screen "分段捻缩" 1280x740, template "模板_设置"
   on GenerateScreen: "TitleUpdater"()
   TextField "Text Field_41" at 427,24 size 154x42; Text '分段捻缩'
   TextField "Text Field_48" at 136,126 size 119x56; Text '第一段:'
   TextField "Text Field_49" at 800,124 size 84x56; Text 'mm/s'
   IOField "IO Field_56" at 693,124 size 91x56; FormatPattern 99.9
      ProcessValue <- "ST_VAR_ZhangLi_HMI_r64Velocity_NianSuo_n{0}"
   IOField "IO Field_1" at 257,126 size 94x56; FormatPattern 999
      ProcessValue <- "ST_VAR_ZhangLi_HMI_r64NianDu_NianSuo_Percent_n{0}"
   TextField "Text Field_2" at 349,125 size 117x56; Text '% ～'
   IOField "IO Field_2" at 440,124 size 115x56; FormatPattern 99.9
      ProcessValue <- "ST_VAR_ZhangLi_HMI_r64NianDu_NianSuo_Percent_n{1}"
   TextField "Text Field_3" at 557,124 size 60x56; Text '%,'
   TextField "Text Field_4" at 604,124 size 82x56; Text '速度:'
   IOField "IO Field_3" at 257,194 size 92x56; FormatPattern 9999
      ProcessValue <- "ST_VAR_ZhangLi_HMI_r64NianDu_NianSuo_n{0}"
   IOField "IO Field_4" at 440,190 size 115x56; FormatPattern 9999
      ProcessValue <- "ST_VAR_ZhangLi_HMI_r64NianDu_NianSuo_n{1}"
   TextField "Text Field_5" at 349,194 size 82x56; Text '捻～'
   TextField "Text Field_6" at 558,190 size 82x56; Text '捻'
   TextField "Text Field_1" at 134,279 size 119x56; Text '第二段:'
   TextField "Text Field_7" at 798,277 size 84x56; Text 'mm/s'
   IOField "IO Field_5" at 691,277 size 91x56; FormatPattern 99.9
      ProcessValue <- "ST_VAR_ZhangLi_HMI_r64Velocity_NianSuo_n{1}"
   IOField "IO Field_6" at 255,279 size 94x56; FormatPattern 99.9
      ProcessValue <- "ST_VAR_ZhangLi_HMI_r64NianDu_NianSuo_Percent_n{1}"
   TextField "Text Field_8" at 347,278 size 117x56; Text '% ～'
   IOField "IO Field_7" at 438,277 size 115x56; FormatPattern 99.9
      ProcessValue <- "ST_VAR_ZhangLi_HMI_r64NianDu_NianSuo_Percent_n{2}"
   TextField "Text Field_9" at 555,277 size 60x56; Text '%,'
   TextField "Text Field_10" at 602,277 size 82x56; Text '速度:'
   IOField "IO Field_8" at 255,347 size 92x56; FormatPattern 9999
      ProcessValue <- "ST_VAR_ZhangLi_HMI_r64NianDu_NianSuo_n{1}"
   IOField "IO Field_9" at 438,343 size 115x56; FormatPattern 9999
      ProcessValue <- "ST_VAR_ZhangLi_HMI_r64NianDu_NianSuo_n{2}"
   TextField "Text Field_11" at 347,347 size 82x56; Text '捻～'
   TextField "Text Field_12" at 556,343 size 82x56; Text '捻'
   TextField "Text Field_13" at 133,436 size 119x56; Text '第三段:'
   TextField "Text Field_14" at 797,434 size 84x56; Text 'mm/s'
   IOField "IO Field_10" at 690,434 size 91x56; FormatPattern 99.9
      ProcessValue <- "ST_VAR_ZhangLi_HMI_r64Velocity_NianSuo_n{2}"
   IOField "IO Field_11" at 254,436 size 94x56; FormatPattern 99.9
      ProcessValue <- "ST_VAR_ZhangLi_HMI_r64NianDu_NianSuo_Percent_n{2}"
   TextField "Text Field_15" at 346,435 size 117x56; Text '% ～'
   IOField "IO Field_12" at 437,434 size 115x56; FormatPattern 999.9
      ProcessValue <- "ST_VAR_ZhangLi_HMI_r64NianDu_NianSuo_Percent_n{3}"
   TextField "Text Field_16" at 554,434 size 60x56; Text '%,'
   TextField "Text Field_17" at 601,434 size 82x56; Text '速度:'
   IOField "IO Field_13" at 254,504 size 92x56; FormatPattern 9999
      ProcessValue <- "ST_VAR_ZhangLi_HMI_r64NianDu_NianSuo_n{2}"
   IOField "IO Field_14" at 437,500 size 115x56; FormatPattern 9999
      ProcessValue <- "ST_VAR_ZhangLi_HMI_r64NianDu_NianSuo_n{3}"
   TextField "Text Field_18" at 346,504 size 82x56; Text '捻～'
   TextField "Text Field_19" at 555,500 size 82x56; Text '捻'
   Button "OBJECT_16" at 227,590 size 228x68; TextOff '启用/停用分段牵伸 / EXIT'
      on Release: InvertBit("ST_VAR_ZhangLi_HMI_bo_NiaoSuo_FenDuan")
      Appearance <- "ST_VAR_ZhangLi_HMI_bo_NiaoSuo_FenDuan"
   Button "OBJECT_1" at 529,590 size 177x68; TextOff '参数复位 / EXIT'
      on Release: ResetBit("ST_VAR_ZhangLi_HMI_bo_NiaoSuo_FenDuan_FuWei")
      on Press: SetBit("ST_VAR_ZhangLi_HMI_bo_NiaoSuo_FenDuan_FuWei")
      Appearance <- "ST_VAR_ZhangLi_HMI_bo_NiaoSuo_FenDuan_FuWei"

screen "包芯纱设定" 1280x740, template "模板_设置"
   on GenerateScreen: "TitleUpdater"()
   TextField "Text Field_81" at 292,64 size 196x42; Text '包芯纱设定'
   TextField "Text Field_82" at 190,134 size 129x56; Text '包芯纱:'
   TextField "Text Field_84" at 190,208 size 210x56; Text '包芯纱牵伸:'
   IOField "IO Field_47" at 418,211 size 140x56; FormatPattern 9.99
      ProcessValue <- "ST_HMI_Var_HMI_r64_QianShenRatio_LaiKa"
   Button "OBJECT_107" at 366,134 size 104x56; TextOff '启用 / EXIT'
      on Release: SetBit("ST_HMI_Var_HMI_bo_LaiKa_Select")
      Appearance <- "ST_HMI_Var_HMI_bo_LaiKa_Select"
      ObjectEnable <- "ST_Main_Var_g_i16_Disable_Status"
   Button "OBJECT_1" at 499,134 size 104x56; TextOff '停用 / EXIT'
      on Release: ResetBit("ST_HMI_Var_HMI_bo_LaiKa_Select")
      Appearance <- "ST_HMI_Var_HMI_bo_LaiKa_Select"
      ObjectEnable <- "ST_Main_Var_g_i16_Disable_Status"
   TextField "文本域_1" at 152,370 size 476x140; Text '说明： 包芯纱只有在“去使能”模式 下，才可“启用”或“停用”。'
   Button "OBJECT_106" at 787,64 size 237x42; TextOff '手动 / EXIT'; TextList "mode_enabled_1"
      ProcessValue <- "ST_Main_Var_g_i16_Mode_Enabled"
      Appearance <- "ST_Main_Var_g_i16_Mode_Enabled"
   Button "OBJECT_5" at 846,254 size 119x60; TextOff '手 动 / EXIT'
      on Release: ResetBit("ST_HMI_Var_HMI_bo_Manual")
      on Press: SetBit("ST_HMI_Var_HMI_bo_Manual")
      Appearance <- "ST_Main_Var_g_i16_Manual_Status"
   Button "OBJECT_6" at 846,150 size 119x60; TextOff '去使能 / EXIT'
      on Release: ResetBit("ST_HMI_Var_HMI_bo_Disable")
      on Press: SetBit("ST_HMI_Var_HMI_bo_Disable")
      Appearance <- "ST_Main_Var_g_i16_Disable_Status"

VB script "timeConverse"
   '注意：要启动脚本，请按下 <Ctrl><空格>，然后就可以看到各种不同函数。
   '通过使用系统函数或 WinCC flexible 对象模型来编写脚本。您可以通过 HMI 运行系统对象很容易地访问系统
   '。挑选对象引用的一个很便利的
   '方式是按下 <Alt><右箭头>。通过使用编程语言 VBScript 的基本功能部件
   '来设计复杂的脚本，并可以直接通过名称，例如 tag = 5，来访问变量。
   'SmartTags("VBS_time_all_hour") = SmartTags("D435_ST_Maintenance_g_r64_Time_All")/3600 
   
   Dim a,b,c,d,e,f
   
   a = SmartTags("ST_Maintenance_g_r64_Time_All(1)")/31536000
   SmartTags("VBS_time_year")=Int(a)
   
   
   b = (a - Int(a))*365
   SmartTags("VBS_time_day")=Int(b)
   
   c =( b - Int(b))*24 
   SmartTags("VBS_time_hour")=Int(c) 
   
   d = (c - Int(c))*60
   SmartTags("VBS_time_min")=Int(d)
   
   e = (d - Int(d))*60
   SmartTags("VBS_time_sec") = Int(e)
    
      
   'SmartTags("VBS_date1") = DateDiff("s", SmartTags("D435_ST_Main_Var_g_dateAndTime0"),Now)
   'SmartTags("VBS_runningRate")= SmartTags("D435_ST_Maintenance_g_r64_Time_All")  / SmartTags("VBS_date1") *100

VB script "TitleUpdater"
   Dim title
   Set title = HmiRuntime.Screens(0).ScreenItems("画面标题")
   title.Text = HmiRuntime.BaseScreenName

VB script "Shasui"
   '注意：要启动脚本，请按下 <Ctrl><空格>，然后就可以看到各种不同函数。
   '通过使用系统函数或 WinCC flexible 对象模型来编写脚本。您可以通过 HMI 运行系统对象很容易地访问系统
   '。挑选对象引用的一个很便利的
   '方式是按下 <Alt><右箭头>。通过使用编程语言 VBScript 的基本功能部件
   '来设计复杂的脚本，并可以直接通过名称，例如 tag = 5，来访问变量。
   
   Dim a
   a=CDbl(SmartTags("ST_Main_Var_g_u16_N_Cycle_Single(1)")) 
   If a<= SmartTags("ST_FC_Var_g_ND") Then 
   	SmartTags("VBS_hengsi_status0")=Int(a/SmartTags("ST_FC_Var_g_ND")*25)
   	SmartTags("VBS_hengsi_status1")=80
   Else
   	SmartTags("VBS_hengsi_status1")=Int((a-SmartTags("ST_FC_Var_g_ND"))/(SmartTags("ST_FC_Var_g_N")-SmartTags("ST_FC_Var_g_ND"))*43)
   	SmartTags("VBS_hengsi_status0")=30
   	
   End If
   
   If SmartTags("ST_Main_Var_g_i16_Mode_Enabled")=512  Then 
   	SmartTags("VBS_hengsi_status1")=80
   	SmartTags("VBS_hengsi_status0")=30
   End If

scheduled task "Job_1"
   on Action: function_f41c6f6c("user_name")

scheduled task "作业_3"
   on Action: ResetBit("VBS_alwaysFalse")
   Triggers <- "1 h"

scheduled task "Task_1"
   on Action: "Shasui"()
   Triggers <- "1 min"

scheduled task "Task_2"
   on Action: "timeConverse"()
   Triggers <- "1 min"
*)